// TIA Portal project "SMS-ENLAB-01-003-1501-001-PLC_V13_SP1_2_V17" (V17) (continued)
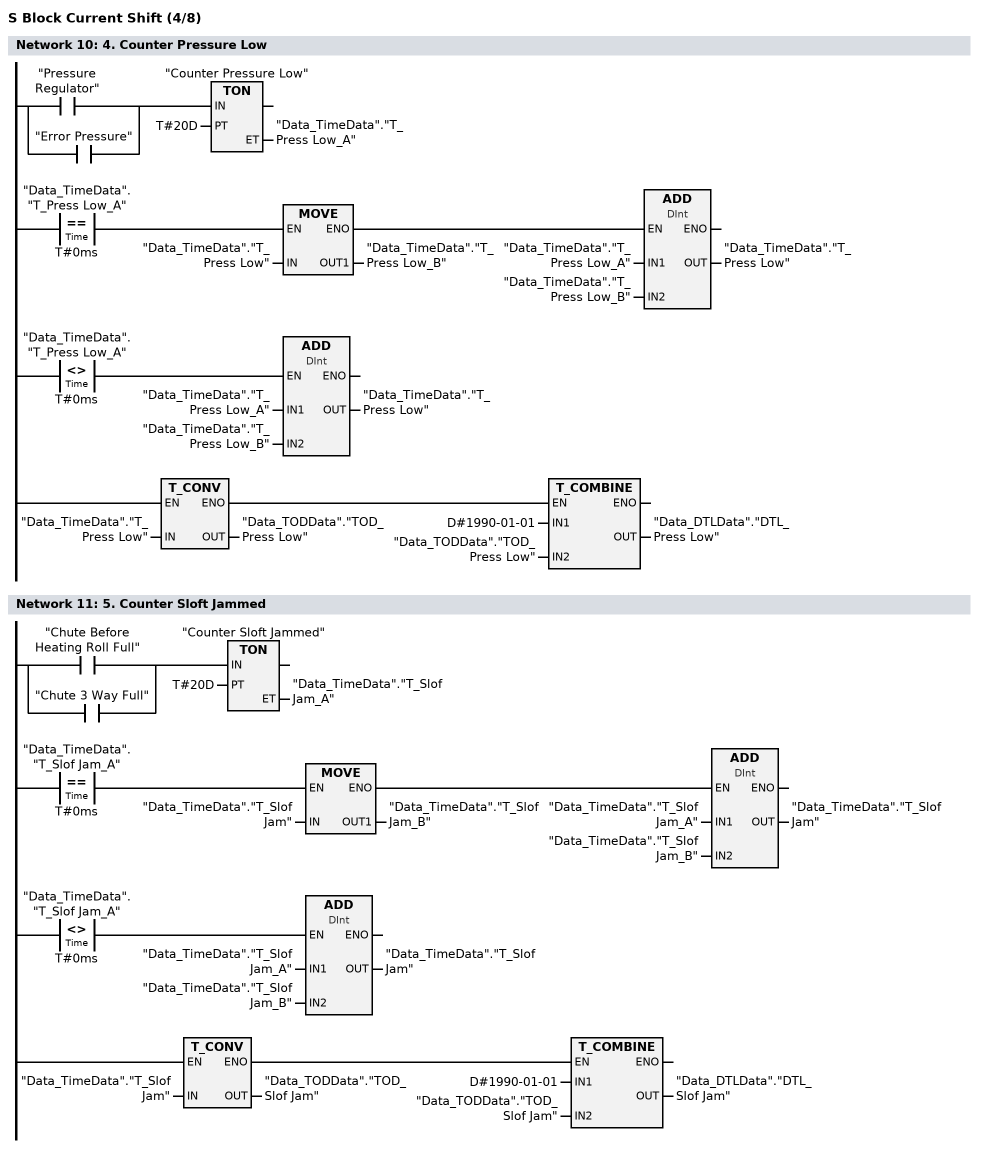
   // ENO of a box is taken as its EN; it also drops when the box reports an error
   "Counter Pressure Low".TON(IN := "Pressure Regulator" OR "Error Pressure",
                           PT := T#20D,
                           ET => "Data_TimeData"."T_Press Low_A");
   IF "Data_TimeData"."T_Press Low_A" = T#0ms THEN
       "Data_TimeData"."T_Press Low_B" := "Data_TimeData"."T_Press Low";
       "Data_TimeData"."T_Press Low" := "Data_TimeData"."T_Press Low_A" + "Data_TimeData"."T_Press Low_B";
   END_IF;
   IF "Data_TimeData"."T_Press Low_A" <> T#0ms THEN
       "Data_TimeData"."T_Press Low" := "Data_TimeData"."T_Press Low_A" + "Data_TimeData"."T_Press Low_B";
   END_IF;
   "Data_TODData"."TOD_Press Low" := T_CONV(IN := "Data_TimeData"."T_Press Low");
   "Data_DTLData"."DTL_Press Low" := T_COMBINE(IN1 := D#1990-01-01, IN2 := "Data_TODData"."TOD_Press Low");
END_REGION

REGION Network 11: 5. Counter Sloft Jammed
   // ENO of a box is taken as its EN; it also drops when the box reports an error
   "Counter Sloft Jammed".TON(IN := "Chute Before Heating Roll Full" OR "Chute 3 Way Full",
                           PT := T#20D,
                           ET => "Data_TimeData"."T_Slof Jam_A");
   IF "Data_TimeData"."T_Slof Jam_A" = T#0ms THEN
       "Data_TimeData"."T_Slof Jam_B" := "Data_TimeData"."T_Slof Jam";
       "Data_TimeData"."T_Slof Jam" := "Data_TimeData"."T_Slof Jam_A" + "Data_TimeData"."T_Slof Jam_B";
   END_IF;
   IF "Data_TimeData"."T_Slof Jam_A" <> T#0ms THEN
       "Data_TimeData"."T_Slof Jam" := "Data_TimeData"."T_Slof Jam_A" + "Data_TimeData"."T_Slof Jam_B";
   END_IF;
   "Data_TODData"."TOD_Slof Jam" := T_CONV(IN := "Data_TimeData"."T_Slof Jam");
   "Data_DTLData"."DTL_Slof Jam" := T_COMBINE(IN1 := D#1990-01-01, IN2 := "Data_TODData"."TOD_Slof Jam");
END_REGION

REGION Network 12: 7. Counter RS Pneumatic Error
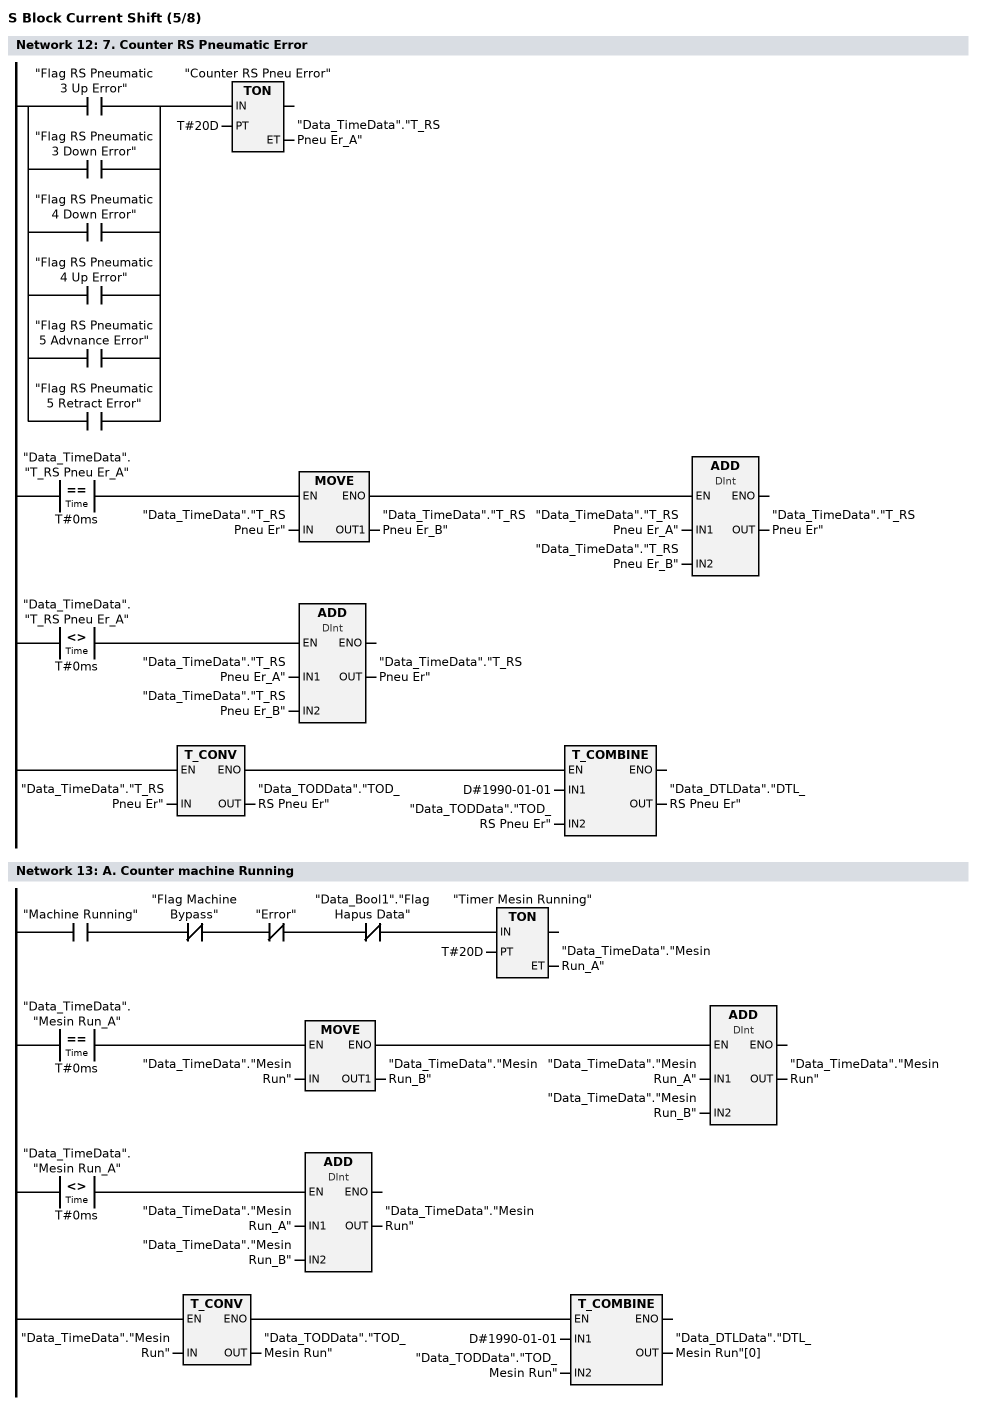
   // ENO of a box is taken as its EN; it also drops when the box reports an error
   "Counter RS Pneu Error".TON(IN := "Flag RS Pneumatic 3 Up Error" OR "Flag RS Pneumatic 3 Down Error" OR "Flag RS Pneumatic 4 Down Error" OR "Flag RS Pneumatic 4 Up Error" OR "Flag RS Pneumatic 5 Advnance Error" OR "Flag RS Pneumatic 5 Retract Error",
                           PT := T#20D,
                           ET => "Data_TimeData"."T_RS Pneu Er_A");
   IF "Data_TimeData"."T_RS Pneu Er_A" = T#0ms THEN
       "Data_TimeData"."T_RS Pneu Er_B" := "Data_TimeData"."T_RS Pneu Er";
       "Data_TimeData"."T_RS Pneu Er" := "Data_TimeData"."T_RS Pneu Er_A" + "Data_TimeData"."T_RS Pneu Er_B";
   END_IF;
   IF "Data_TimeData"."T_RS Pneu Er_A" <> T#0ms THEN
       "Data_TimeData"."T_RS Pneu Er" := "Data_TimeData"."T_RS Pneu Er_A" + "Data_TimeData"."T_RS Pneu Er_B";
   END_IF;
   "Data_TODData"."TOD_RS Pneu Er" := T_CONV(IN := "Data_TimeData"."T_RS Pneu Er");
   "Data_DTLData"."DTL_RS Pneu Er" := T_COMBINE(IN1 := D#1990-01-01, IN2 := "Data_TODData"."TOD_RS Pneu Er");
END_REGION

REGION Network 13: A. Counter machine Running
   // ENO of a box is taken as its EN; it also drops when the box reports an error
   "Timer Mesin Running".TON(IN := "Machine Running" AND NOT "Flag Machine Bypass" AND NOT "Error" AND NOT "Data_Bool1"."Flag Hapus Data",
                           PT := T#20D,
                           ET => "Data_TimeData"."Mesin Run_A");
   IF "Data_TimeData"."Mesin Run_A" = T#0ms THEN
       "Data_TimeData"."Mesin Run_B" := "Data_TimeData"."Mesin Run";
       "Data_TimeData"."Mesin Run" := "Data_TimeData"."Mesin Run_A" + "Data_TimeData"."Mesin Run_B";
   END_IF;
   IF "Data_TimeData"."Mesin Run_A" <> T#0ms THEN
       "Data_TimeData"."Mesin Run" := "Data_TimeData"."Mesin Run_A" + "Data_TimeData"."Mesin Run_B";
   END_IF;
   "Data_TODData"."TOD_Mesin Run" := T_CONV(IN := "Data_TimeData"."Mesin Run");
   "Data_DTLData"."DTL_Mesin Run"[0] := T_COMBINE(IN1 := D#1990-01-01, IN2 := "Data_TODData"."TOD_Mesin Run");
END_REGION

REGION Network 14: B. Counter machine Running Baypass Stamp
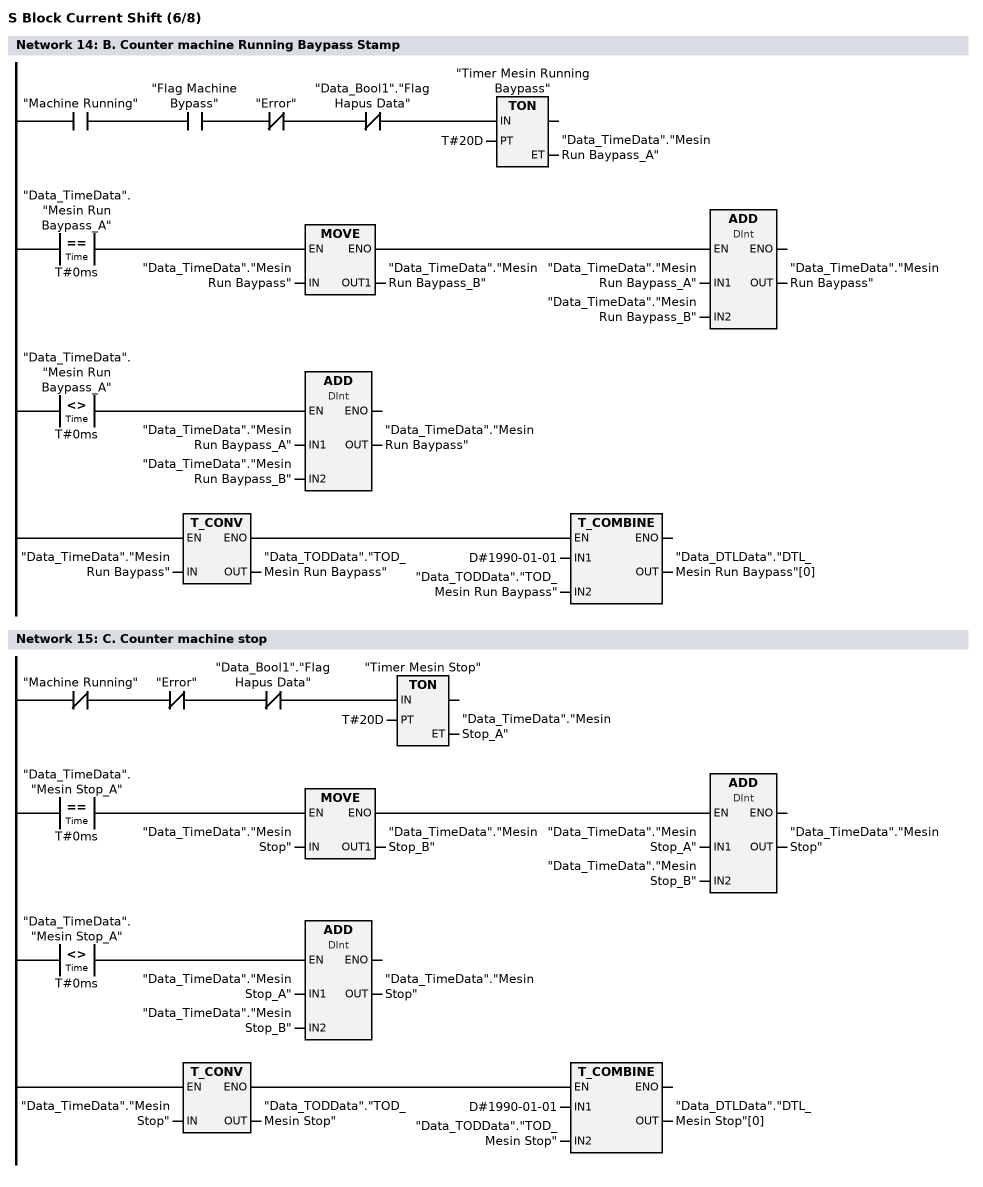
   // ENO of a box is taken as its EN; it also drops when the box reports an error
   "Timer Mesin Running Baypass".TON(IN := "Machine Running" AND "Flag Machine Bypass" AND NOT "Error" AND NOT "Data_Bool1"."Flag Hapus Data",
                           PT := T#20D,
                           ET => "Data_TimeData"."Mesin Run Baypass_A");
   IF "Data_TimeData"."Mesin Run Baypass_A" = T#0ms THEN
       "Data_TimeData"."Mesin Run Baypass_B" := "Data_TimeData"."Mesin Run Baypass";
       "Data_TimeData"."Mesin Run Baypass" := "Data_TimeData"."Mesin Run Baypass_A" + "Data_TimeData"."Mesin Run Baypass_B";
   END_IF;
   IF "Data_TimeData"."Mesin Run Baypass_A" <> T#0ms THEN
       "Data_TimeData"."Mesin Run Baypass" := "Data_TimeData"."Mesin Run Baypass_A" + "Data_TimeData"."Mesin Run Baypass_B";
   END_IF;
   "Data_TODData"."TOD_Mesin Run Baypass" := T_CONV(IN := "Data_TimeData"."Mesin Run Baypass");
   "Data_DTLData"."DTL_Mesin Run Baypass"[0] := T_COMBINE(IN1 := D#1990-01-01,
                           IN2 := "Data_TODData"."TOD_Mesin Run Baypass");
END_REGION

REGION Network 15: C. Counter machine stop
   // ENO of a box is taken as its EN; it also drops when the box reports an error
   "Timer Mesin Stop".TON(IN := NOT "Machine Running" AND NOT "Error" AND NOT "Data_Bool1"."Flag Hapus Data",
                          PT := T#20D,
                          ET => "Data_TimeData"."Mesin Stop_A");
   IF "Data_TimeData"."Mesin Stop_A" = T#0ms THEN
       "Data_TimeData"."Mesin Stop_B" := "Data_TimeData"."Mesin Stop";
       "Data_TimeData"."Mesin Stop" := "Data_TimeData"."Mesin Stop_A" + "Data_TimeData"."Mesin Stop_B";
   END_IF;
   IF "Data_TimeData"."Mesin Stop_A" <> T#0ms THEN
       "Data_TimeData"."Mesin Stop" := "Data_TimeData"."Mesin Stop_A" + "Data_TimeData"."Mesin Stop_B";
   END_IF;
   "Data_TODData"."TOD_Mesin Stop" := T_CONV(IN := "Data_TimeData"."Mesin Stop");
   "Data_DTLData"."DTL_Mesin Stop"[0] := T_COMBINE(IN1 := D#1990-01-01, IN2 := "Data_TODData"."TOD_Mesin Stop");
END_REGION

REGION Network 16: D. Counter Machine Error
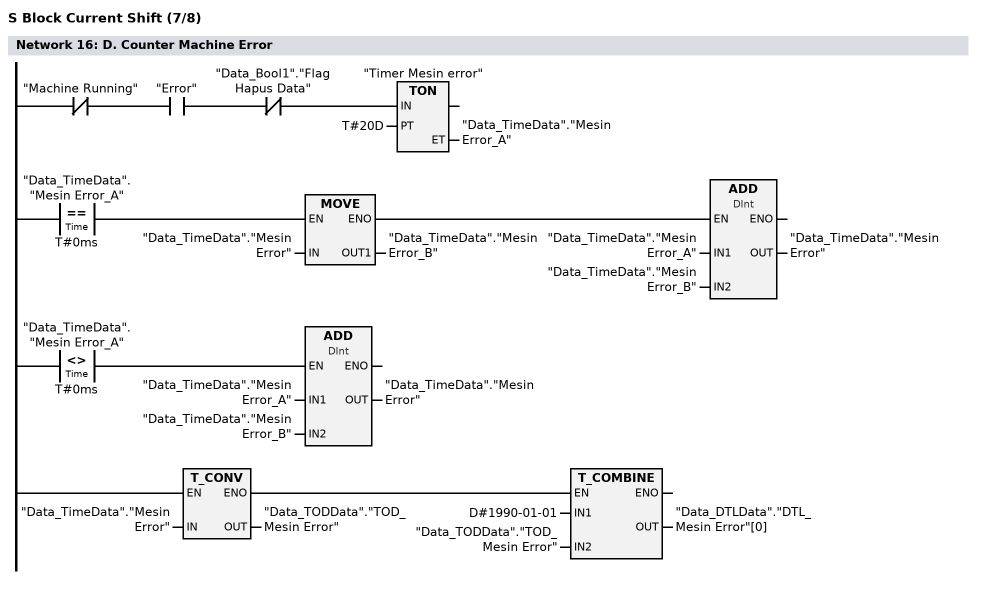
   // ENO of a box is taken as its EN; it also drops when the box reports an error
   "Timer Mesin error".TON(IN := NOT "Machine Running" AND "Error" AND NOT "Data_Bool1"."Flag Hapus Data",
                           PT := T#20D,
                           ET => "Data_TimeData"."Mesin Error_A");
   IF "Data_TimeData"."Mesin Error_A" = T#0ms THEN
       "Data_TimeData"."Mesin Error_B" := "Data_TimeData"."Mesin Error";
       "Data_TimeData"."Mesin Error" := "Data_TimeData"."Mesin Error_A" + "Data_TimeData"."Mesin Error_B";
   END_IF;
   IF "Data_TimeData"."Mesin Error_A" <> T#0ms THEN
       "Data_TimeData"."Mesin Error" := "Data_TimeData"."Mesin Error_A" + "Data_TimeData"."Mesin Error_B";
   END_IF;
   "Data_TODData"."TOD_Mesin Error" := T_CONV(IN := "Data_TimeData"."Mesin Error");
   "Data_DTLData"."DTL_Mesin Error"[0] := T_COMBINE(IN1 := D#1990-01-01,
                           IN2 := "Data_TODData"."TOD_Mesin Error");
END_REGION

REGION Network 17: % Persen Counter Mesin Terhadap Lama Current Shift
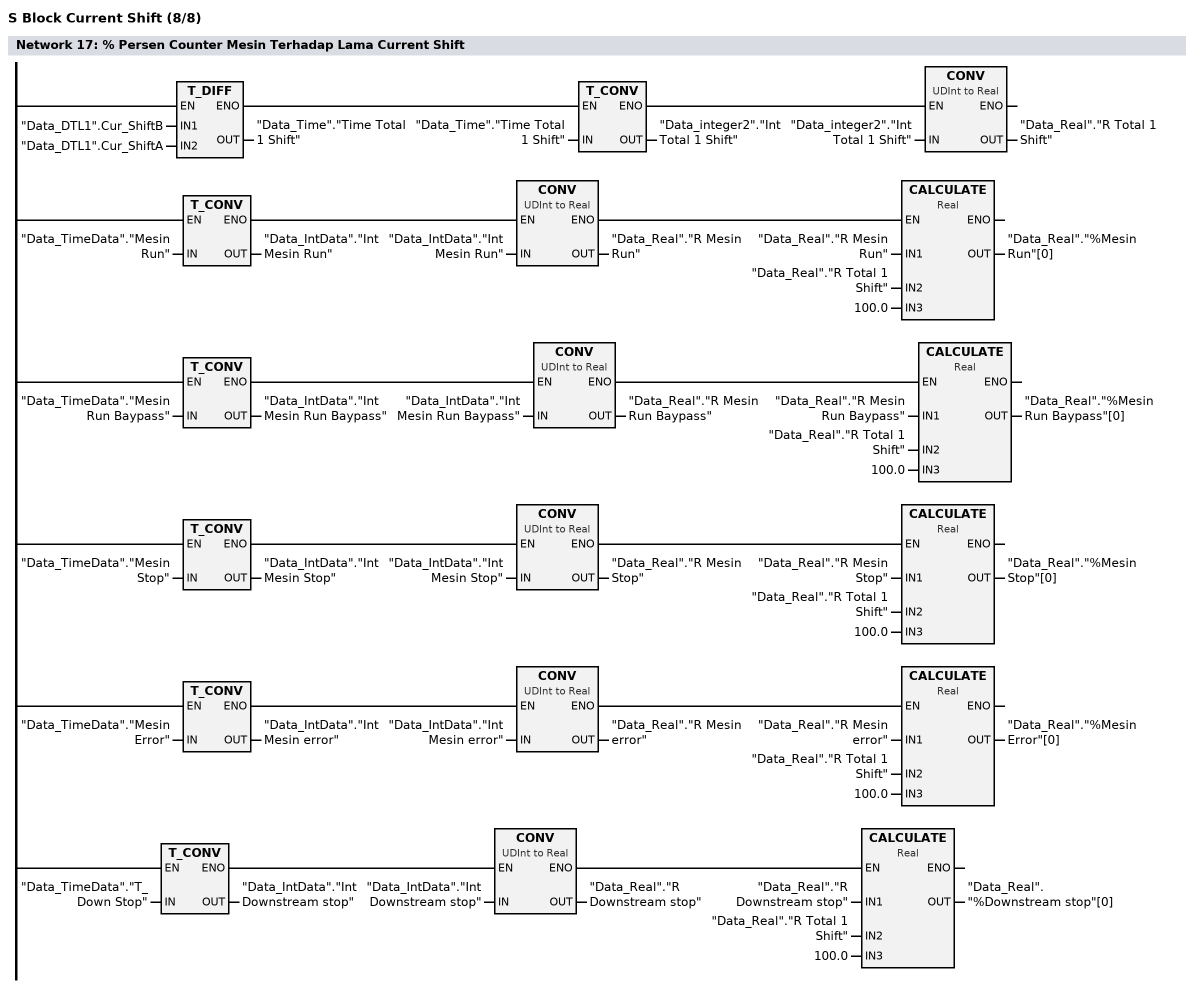
   // ENO of a box is taken as its EN; it also drops when the box reports an error
   "Data_Time"."Time Total 1 Shift" := T_DIFF(IN1 := "Data_DTL1".Cur_ShiftB, IN2 := "Data_DTL1".Cur_ShiftA);
   "Data_integer2"."Int Total 1 Shift" := T_CONV(IN := "Data_Time"."Time Total 1 Shift");
   "Data_Real"."R Total 1 Shift" := UDINT_TO_REAL("Data_integer2"."Int Total 1 Shift");
   "Data_IntData"."Int Mesin Run" := T_CONV(IN := "Data_TimeData"."Mesin Run");
   "Data_Real"."R Mesin Run" := UDINT_TO_REAL("Data_IntData"."Int Mesin Run");
   "Data_Real"."%Mesin Run"[0] := ("Data_Real"."R Mesin Run"/"Data_Real"."R Total 1 Shift")*100.0;
   "Data_IntData"."Int Mesin Run Baypass" := T_CONV(IN := "Data_TimeData"."Mesin Run Baypass");
   "Data_Real"."R Mesin Run Baypass" := UDINT_TO_REAL("Data_IntData"."Int Mesin Run Baypass");
   "Data_Real"."%Mesin Run Baypass"[0] := ("Data_Real"."R Mesin Run Baypass"/"Data_Real"."R Total 1 Shift")*100.0;
   "Data_IntData"."Int Mesin Stop" := T_CONV(IN := "Data_TimeData"."Mesin Stop");
   "Data_Real"."R Mesin Stop" := UDINT_TO_REAL("Data_IntData"."Int Mesin Stop");
   "Data_Real"."%Mesin Stop"[0] := ("Data_Real"."R Mesin Stop"/"Data_Real"."R Total 1 Shift")*100.0;
   "Data_IntData"."Int Mesin error" := T_CONV(IN := "Data_TimeData"."Mesin Error");
   "Data_Real"."R Mesin error" := UDINT_TO_REAL("Data_IntData"."Int Mesin error");
   "Data_Real"."%Mesin Error"[0] := ("Data_Real"."R Mesin error"/"Data_Real"."R Total 1 Shift")*100.0;
   "Data_IntData"."Int Downstream stop" := T_CONV(IN := "Data_TimeData"."T_Down Stop");
   "Data_Real"."R Downstream stop" := UDINT_TO_REAL("Data_IntData"."Int Downstream stop");
   "Data_Real"."%Downstream stop"[0] := ("Data_Real"."R Downstream stop"/"Data_Real"."R Total 1 Shift")*100.0;
END_REGION
END_FUNCTION_BLOCK

FUNCTION_BLOCK "Block Labeling"   // FB5, LAD
{ S7_Optimized_Access := 'TRUE' }
VERSION : 0.1
   VAR_TEMP   // added for the SCL form of the ladder/FBD networks
      _w1 : Bool;
      _w2 : Bool;
      _w3 : Bool;
      _w4 : Bool;
      _w5 : Bool;
   END_VAR
BEGIN

REGION Network 1: By pass ON
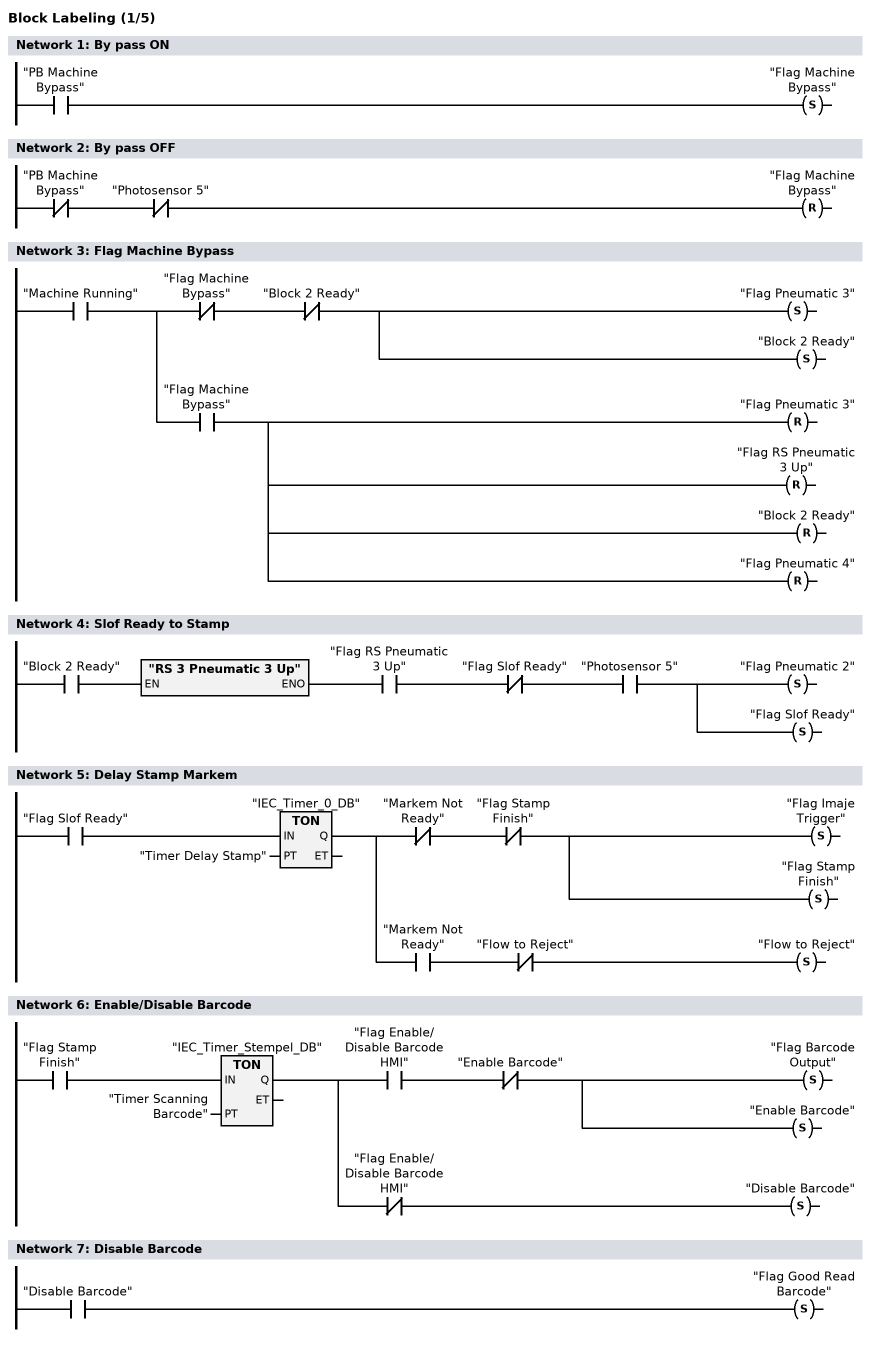
   RUNG wire#powerrail
      Contact( "PB Machine Bypass" )
      S_Coil( "Flag Machine Bypass" )
   END_RUNG
   // the same network as SCL:
   IF "PB Machine Bypass" THEN "Flag Machine Bypass" := TRUE; END_IF;
END_REGION

REGION Network 2: By pass OFF
   RUNG wire#powerrail
      I_Contact( "PB Machine Bypass" )
      I_Contact( "Photosensor 5" )
      R_Coil( "Flag Machine Bypass" )
   END_RUNG
   // the same network as SCL:
   IF NOT "PB Machine Bypass" AND NOT "Photosensor 5" THEN "Flag Machine Bypass" := FALSE; END_IF;
END_REGION

REGION Network 3: Flag Machine Bypass
   RUNG wire#powerrail
      Contact( "Machine Running" )
      wire#w1
      I_Contact( "Flag Machine Bypass" )
      I_Contact( "Block 2 Ready" )
      wire#w2
      S_Coil( "Flag Pneumatic 3" )
   END_RUNG
   RUNG wire#w2
      S_Coil( "Block 2 Ready" )
   END_RUNG
   RUNG wire#w1
      Contact( "Flag Machine Bypass" )
      wire#w3
      R_Coil( "Flag Pneumatic 3" )
   END_RUNG
   RUNG wire#w3
      R_Coil( "Flag RS Pneumatic 3 Up" )
   END_RUNG
   RUNG wire#w3
      R_Coil( "Block 2 Ready" )
   END_RUNG
   RUNG wire#w3
      R_Coil( "Flag Pneumatic 4" )
   END_RUNG
   // the same network as SCL:
   IF "Machine Running" AND NOT "Flag Machine Bypass" AND NOT "Block 2 Ready" THEN
       "Flag Pneumatic 3" := TRUE;
       "Block 2 Ready" := TRUE;
   END_IF;
   IF "Machine Running" AND "Flag Machine Bypass" THEN
       "Flag Pneumatic 3" := FALSE;
       "Flag RS Pneumatic 3 Up" := FALSE;
       "Block 2 Ready" := FALSE;
       "Flag Pneumatic 4" := FALSE;
   END_IF;
END_REGION

REGION Network 4: Slof Ready to Stamp
   RUNG wire#powerrail
      Contact( "Block 2 Ready" )
      "RS 3 Pneumatic 3 Up"()
      Contact( "Flag RS Pneumatic 3 Up" )
      I_Contact( "Flag Slof Ready" )
      Contact( "Photosensor 5" )
      wire#w1
      S_Coil( "Flag Pneumatic 2" )
   END_RUNG
   RUNG wire#w1
      S_Coil( "Flag Slof Ready" )
   END_RUNG
   // the same network as SCL:
   "RS 3 Pneumatic 3 Up"(EN := "Block 2 Ready", ENO => #_w1);
   IF #_w1 AND "Flag RS Pneumatic 3 Up" AND NOT "Flag Slof Ready" AND "Photosensor 5" THEN
       "Flag Pneumatic 2" := TRUE;
       "Flag Slof Ready" := TRUE;
   END_IF;
END_REGION

REGION Network 5: Delay Stamp Markem
   "IEC_Timer_0_DB".TON(IN := "Flag Slof Ready", PT := "Timer Delay Stamp");
   IF "IEC_Timer_0_DB".Q AND NOT "Markem Not Ready" AND NOT "Flag Stamp Finish" THEN
       "Flag Imaje Trigger" := TRUE;
       "Flag Stamp Finish" := TRUE;
   END_IF;
   IF "IEC_Timer_0_DB".Q AND "Markem Not Ready" AND NOT "Flow to Reject" THEN
       "Flow to Reject" := TRUE;
   END_IF;
END_REGION

REGION Network 6: Enable/Disable Barcode
   "IEC_Timer_Stempel_DB".TON(IN := "Flag Stamp Finish", PT := "Timer Scanning Barcode");
   IF "IEC_Timer_Stempel_DB".Q AND "Flag Enable/Disable Barcode HMI" AND NOT "Enable Barcode" THEN
       "Flag Barcode Output" := TRUE;
       "Enable Barcode" := TRUE;
   END_IF;
   IF "IEC_Timer_Stempel_DB".Q AND NOT "Flag Enable/Disable Barcode HMI" THEN
       "Disable Barcode" := TRUE;
   END_IF;
END_REGION

REGION Network 7: Disable Barcode
   RUNG wire#powerrail
      Contact( "Disable Barcode" )
      S_Coil( "Flag Good Read Barcode" )
   END_RUNG
   // the same network as SCL:
   IF "Disable Barcode" THEN "Flag Good Read Barcode" := TRUE; END_IF;
END_REGION

REGION Network 8: Check Barcode
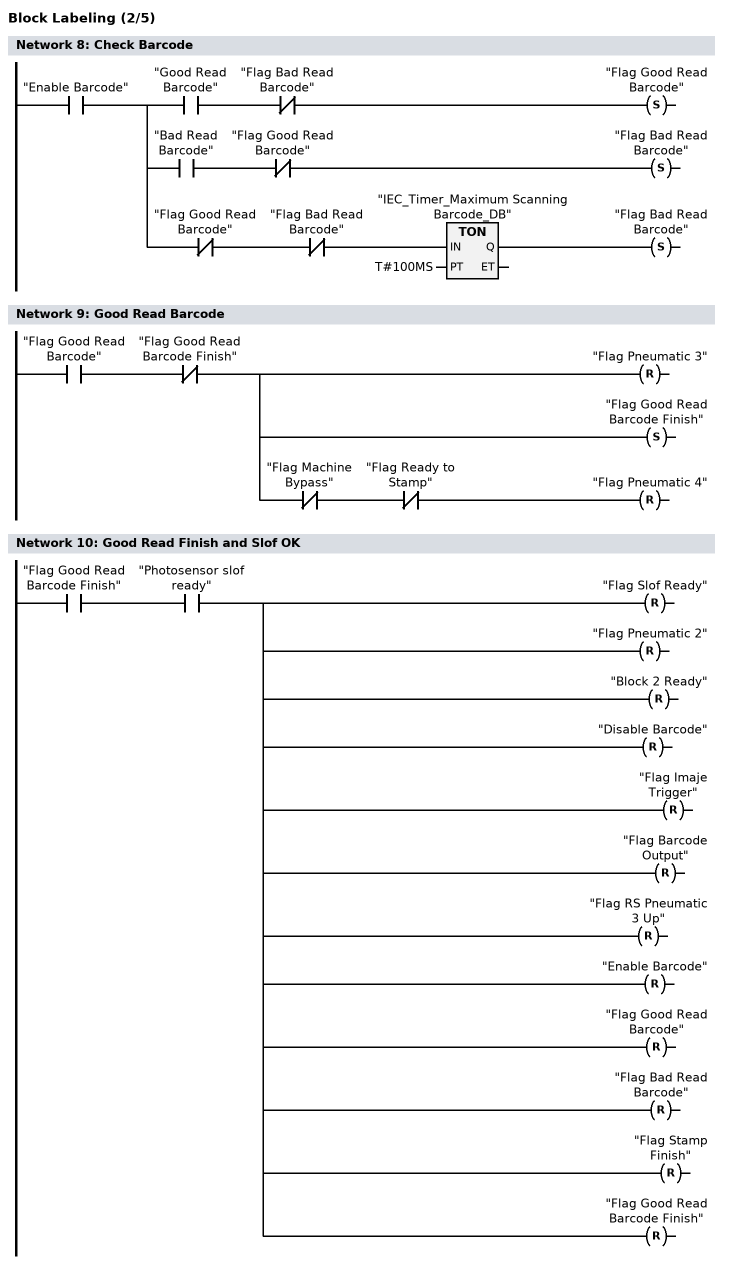
   IF "Enable Barcode" AND "Good Read Barcode" AND NOT "Flag Bad Read Barcode" THEN
       "Flag Good Read Barcode" := TRUE;
   END_IF;
   IF "Enable Barcode" AND "Bad Read Barcode" AND NOT "Flag Good Read Barcode" THEN
       "Flag Bad Read Barcode" := TRUE;
   END_IF;
   "IEC_Timer_Maximum Scanning Barcode_DB".TON(IN := "Enable Barcode" AND NOT "Flag Good Read Barcode" AND NOT "Flag Bad Read Barcode",
                           PT := T#100MS);
   IF "IEC_Timer_Maximum Scanning Barcode_DB".Q THEN "Flag Bad Read Barcode" := TRUE; END_IF;
END_REGION

REGION Network 9: Good Read Barcode
   RUNG wire#powerrail
      Contact( "Flag Good Read Barcode" )
      I_Contact( "Flag Good Read Barcode Finish" )
      wire#w1
      R_Coil( "Flag Pneumatic 3" )
   END_RUNG
   RUNG wire#w1
      S_Coil( "Flag Good Read Barcode Finish" )
   END_RUNG
   RUNG wire#w1
      I_Contact( "Flag Machine Bypass" )
      I_Contact( "Flag Ready to Stamp" )
      R_Coil( "Flag Pneumatic 4" )
   END_RUNG
   // the same network as SCL:
   #_w1 := "Flag Good Read Barcode" AND NOT "Flag Good Read Barcode Finish";
   IF #_w1 THEN
       "Flag Pneumatic 3" := FALSE;
       "Flag Good Read Barcode Finish" := TRUE;
   END_IF;
   IF #_w1 AND NOT "Flag Machine Bypass" AND NOT "Flag Ready to Stamp" THEN
       "Flag Pneumatic 4" := FALSE;
   END_IF;
END_REGION

REGION Network 10: Good Read Finish and Slof OK
   RUNG wire#powerrail
      Contact( "Flag Good Read Barcode Finish" )
      Contact( "Photosensor slof ready" )
      wire#w1
      R_Coil( "Flag Slof Ready" )
   END_RUNG
   RUNG wire#w1
      R_Coil( "Flag Pneumatic 2" )
   END_RUNG
   RUNG wire#w1
      R_Coil( "Block 2 Ready" )
   END_RUNG
   RUNG wire#w1
      R_Coil( "Disable Barcode" )
   END_RUNG
   RUNG wire#w1
      R_Coil( "Flag Imaje Trigger" )
   END_RUNG
   RUNG wire#w1
      R_Coil( "Flag Barcode Output" )
   END_RUNG
   RUNG wire#w1
      R_Coil( "Flag RS Pneumatic 3 Up" )
   END_RUNG
   RUNG wire#w1
      R_Coil( "Enable Barcode" )
   END_RUNG
   RUNG wire#w1
      R_Coil( "Flag Good Read Barcode" )
   END_RUNG
   RUNG wire#w1
      R_Coil( "Flag Bad Read Barcode" )
   END_RUNG
   RUNG wire#w1
      R_Coil( "Flag Stamp Finish" )
   END_RUNG
   RUNG wire#w1
      R_Coil( "Flag Good Read Barcode Finish" )
   END_RUNG
   // the same network as SCL:
   IF "Flag Good Read Barcode Finish" AND "Photosensor slof ready" THEN
       "Flag Slof Ready" := FALSE;
       "Flag Pneumatic 2" := FALSE;
       "Block 2 Ready" := FALSE;
       "Disable Barcode" := FALSE;
       "Flag Imaje Trigger" := FALSE;
       "Flag Barcode Output" := FALSE;
       "Flag RS Pneumatic 3 Up" := FALSE;
       "Enable Barcode" := FALSE;
       "Flag Good Read Barcode" := FALSE;
       "Flag Bad Read Barcode" := FALSE;
       "Flag Stamp Finish" := FALSE;
       "Flag Good Read Barcode Finish" := FALSE;
   END_IF;
END_REGION

REGION Network 11: Set Section Reject
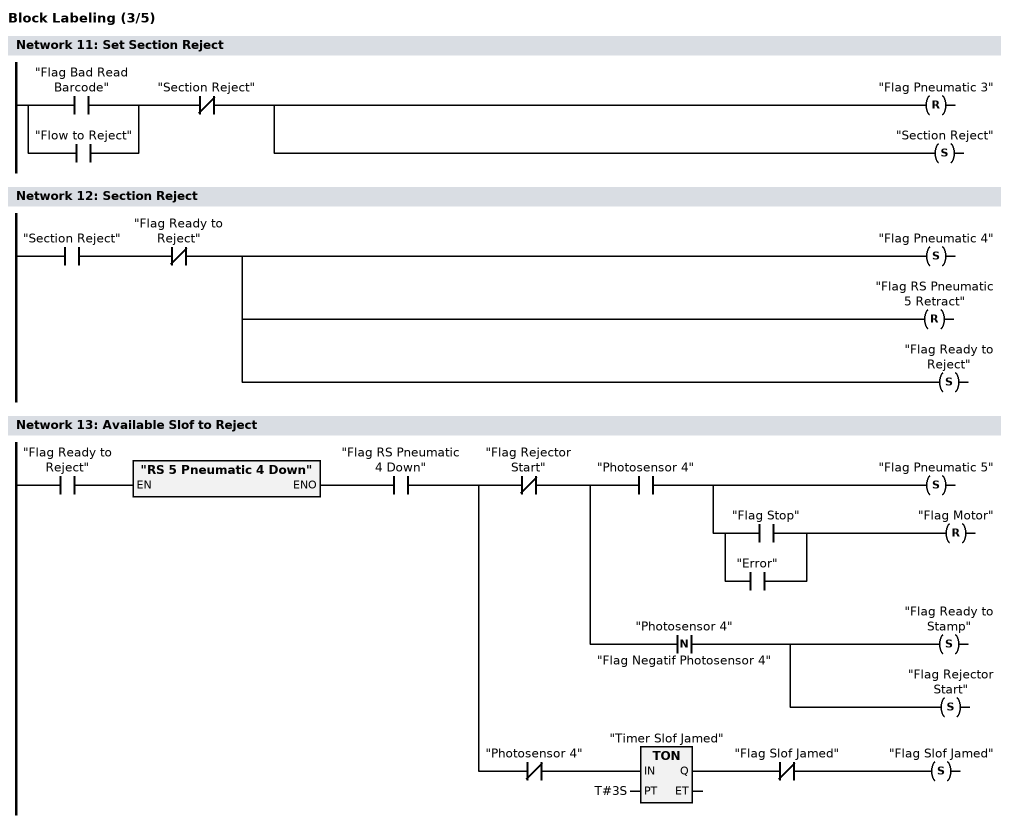
   RUNG wire#powerrail
      Contact( "Flag Bad Read Barcode" )
      wire#w1
      I_Contact( "Section Reject" )
      wire#w2
      R_Coil( "Flag Pneumatic 3" )
   END_RUNG
   RUNG wire#powerrail
      Contact( "Flow to Reject" )
   END_RUNG wire#w1
   RUNG wire#w2
      S_Coil( "Section Reject" )
   END_RUNG
   // the same network as SCL:
   IF ("Flag Bad Read Barcode" OR "Flow to Reject") AND NOT "Section Reject" THEN
       "Flag Pneumatic 3" := FALSE;
       "Section Reject" := TRUE;
   END_IF;
END_REGION

REGION Network 12: Section Reject
   RUNG wire#powerrail
      Contact( "Section Reject" )
      I_Contact( "Flag Ready to Reject" )
      wire#w1
      S_Coil( "Flag Pneumatic 4" )
   END_RUNG
   RUNG wire#w1
      R_Coil( "Flag RS Pneumatic 5 Retract" )
   END_RUNG
   RUNG wire#w1
      S_Coil( "Flag Ready to Reject" )
   END_RUNG
   // the same network as SCL:
   IF "Section Reject" AND NOT "Flag Ready to Reject" THEN
       "Flag Pneumatic 4" := TRUE;
       "Flag RS Pneumatic 5 Retract" := FALSE;
       "Flag Ready to Reject" := TRUE;
   END_IF;
END_REGION

REGION Network 13: Available Slof to Reject
   "RS 5 Pneumatic 4 Down"(EN := "Flag Ready to Reject", ENO => #_w1);
   #_w2 := #_w1 AND "Flag RS Pneumatic 4 Down";
   #_w3 := #_w2 AND NOT "Flag Rejector Start";
   #_w4 := #_w3 AND "Photosensor 4";
   IF #_w4 THEN "Flag Pneumatic 5" := TRUE; END_IF;
   IF #_w4 AND ("Flag Stop" OR "Error") THEN "Flag Motor" := FALSE; END_IF;
   #_w5 := #_w3 AND NOT "Photosensor 4" AND "Flag Negatif Photosensor 4";   // falling edge of "Photosensor 4"
   "Flag Negatif Photosensor 4" := "Photosensor 4";
   IF #_w5 THEN
       "Flag Ready to Stamp" := TRUE;
       "Flag Rejector Start" := TRUE;
   END_IF;
   "Timer Slof Jamed".TON(IN := #_w2 AND NOT "Photosensor 4", PT := T#3S);
   IF "Timer Slof Jamed".Q AND NOT "Flag Slof Jamed" THEN "Flag Slof Jamed" := TRUE; END_IF;
END_REGION

REGION Network 14: Ready to Stamp again
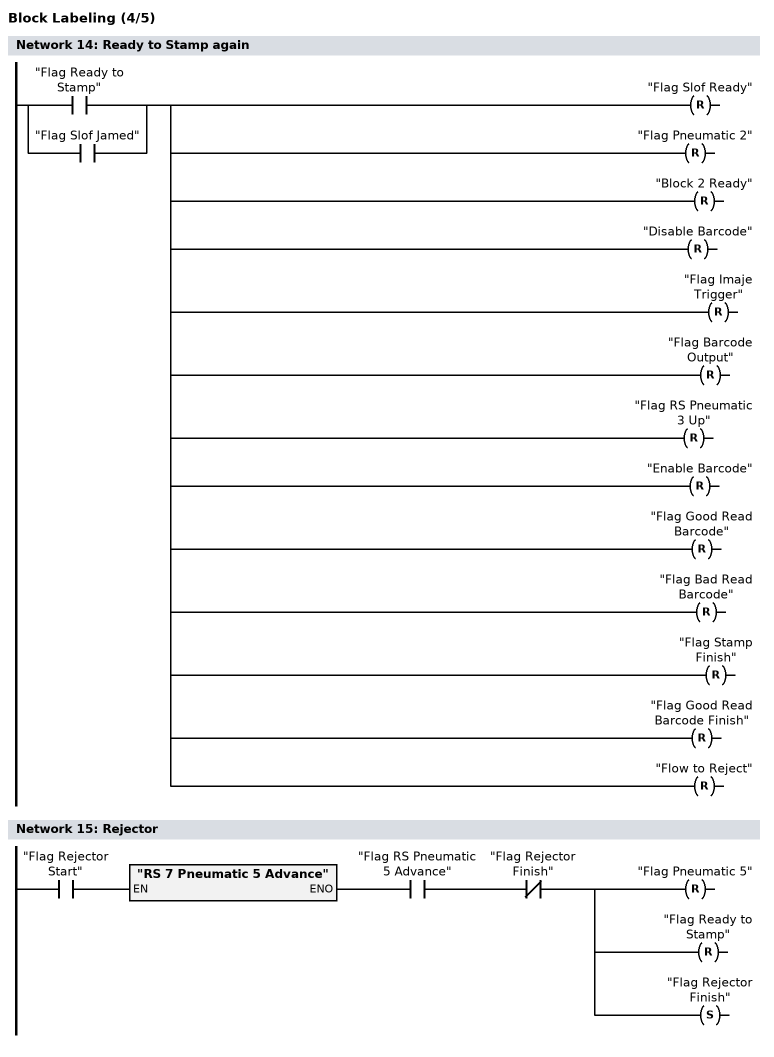
   RUNG wire#powerrail
      Contact( "Flag Ready to Stamp" )
      wire#w1
      R_Coil( "Flag Slof Ready" )
   END_RUNG
   RUNG wire#powerrail
      Contact( "Flag Slof Jamed" )
   END_RUNG wire#w1
   RUNG wire#w1
      R_Coil( "Flag Pneumatic 2" )
   END_RUNG
   RUNG wire#w1
      R_Coil( "Block 2 Ready" )
   END_RUNG
   RUNG wire#w1
      R_Coil( "Disable Barcode" )
   END_RUNG
   RUNG wire#w1
      R_Coil( "Flag Imaje Trigger" )
   END_RUNG
   RUNG wire#w1
      R_Coil( "Flag Barcode Output" )
   END_RUNG
   RUNG wire#w1
      R_Coil( "Flag RS Pneumatic 3 Up" )
   END_RUNG
   RUNG wire#w1
      R_Coil( "Enable Barcode" )
   END_RUNG
   RUNG wire#w1
      R_Coil( "Flag Good Read Barcode" )
   END_RUNG
   RUNG wire#w1
      R_Coil( "Flag Bad Read Barcode" )
   END_RUNG
   RUNG wire#w1
      R_Coil( "Flag Stamp Finish" )
   END_RUNG
   RUNG wire#w1
      R_Coil( "Flag Good Read Barcode Finish" )
   END_RUNG
   RUNG wire#w1
      R_Coil( "Flow to Reject" )
   END_RUNG
   // the same network as SCL:
   IF "Flag Ready to Stamp" OR "Flag Slof Jamed" THEN
       "Flag Slof Ready" := FALSE;
       "Flag Pneumatic 2" := FALSE;
       "Block 2 Ready" := FALSE;
       "Disable Barcode" := FALSE;
       "Flag Imaje Trigger" := FALSE;
       "Flag Barcode Output" := FALSE;
       "Flag RS Pneumatic 3 Up" := FALSE;
       "Enable Barcode" := FALSE;
       "Flag Good Read Barcode" := FALSE;
       "Flag Bad Read Barcode" := FALSE;
       "Flag Stamp Finish" := FALSE;
       "Flag Good Read Barcode Finish" := FALSE;
       "Flow to Reject" := FALSE;
   END_IF;
END_REGION

REGION Network 15: Rejector
   RUNG wire#powerrail
      Contact( "Flag Rejector Start" )
      "RS 7 Pneumatic 5 Advance"()
      Contact( "Flag RS Pneumatic 5 Advance" )
      I_Contact( "Flag Rejector Finish" )
      wire#w1
      R_Coil( "Flag Pneumatic 5" )
   END_RUNG
   RUNG wire#w1
      R_Coil( "Flag Ready to Stamp" )
   END_RUNG
   RUNG wire#w1
      S_Coil( "Flag Rejector Finish" )
   END_RUNG
   // the same network as SCL:
   "RS 7 Pneumatic 5 Advance"(EN := "Flag Rejector Start", ENO => #_w1);
   IF #_w1 AND "Flag RS Pneumatic 5 Advance" AND NOT "Flag Rejector Finish" THEN
       "Flag Pneumatic 5" := FALSE;
       "Flag Ready to Stamp" := FALSE;
       "Flag Rejector Finish" := TRUE;
   END_IF;
END_REGION

REGION Network 16: Rejector Finish
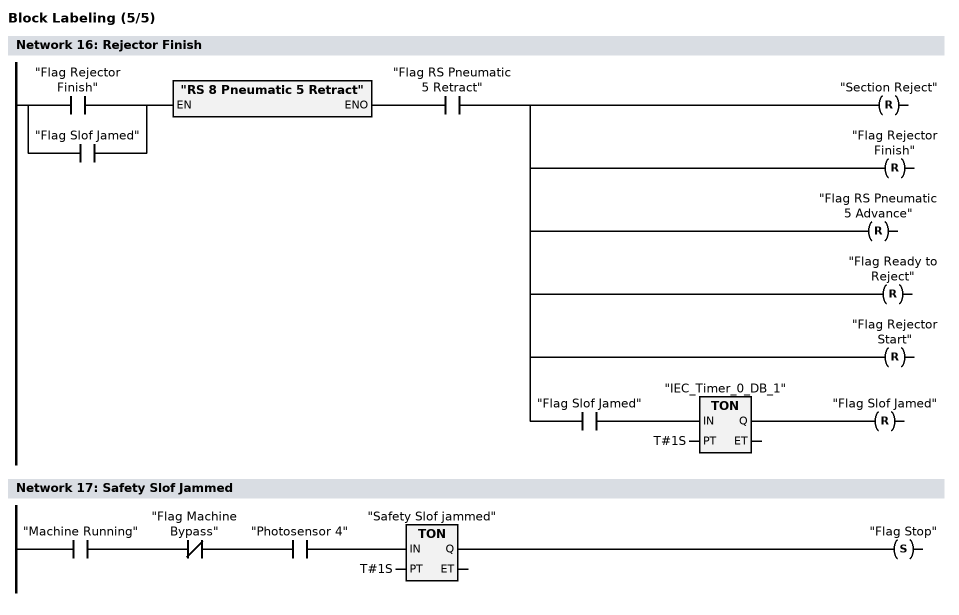
   "RS 8 Pneumatic 5 Retract"(EN := "Flag Rejector Finish" OR "Flag Slof Jamed", ENO => #_w1);
   #_w2 := #_w1 AND "Flag RS Pneumatic 5 Retract";
   IF #_w2 THEN
       "Section Reject" := FALSE;
       "Flag Rejector Finish" := FALSE;
       "Flag RS Pneumatic 5 Advance" := FALSE;
       "Flag Ready to Reject" := FALSE;
       "Flag Rejector Start" := FALSE;
   END_IF;
   "IEC_Timer_0_DB_1".TON(IN := #_w2 AND "Flag Slof Jamed", PT := T#1S);
   IF "IEC_Timer_0_DB_1".Q THEN "Flag Slof Jamed" := FALSE; END_IF;
END_REGION

REGION Network 17: Safety Slof Jammed
   "Safety Slof jammed".TON(IN := "Machine Running" AND NOT "Flag Machine Bypass" AND "Photosensor 4",
                           PT := T#1S);
   IF "Safety Slof jammed".Q THEN "Flag Stop" := TRUE; END_IF;
END_REGION
END_FUNCTION_BLOCK

FUNCTION_BLOCK "Block Focke"   // FB6, LAD
{ S7_Optimized_Access := 'TRUE' }
VERSION : 0.1
   VAR_TEMP   // added for the SCL form of the ladder/FBD networks
      _w1 : Bool;
   END_VAR
BEGIN

REGION Network 1: Enable/Disable Error Chute Before Heating Roll
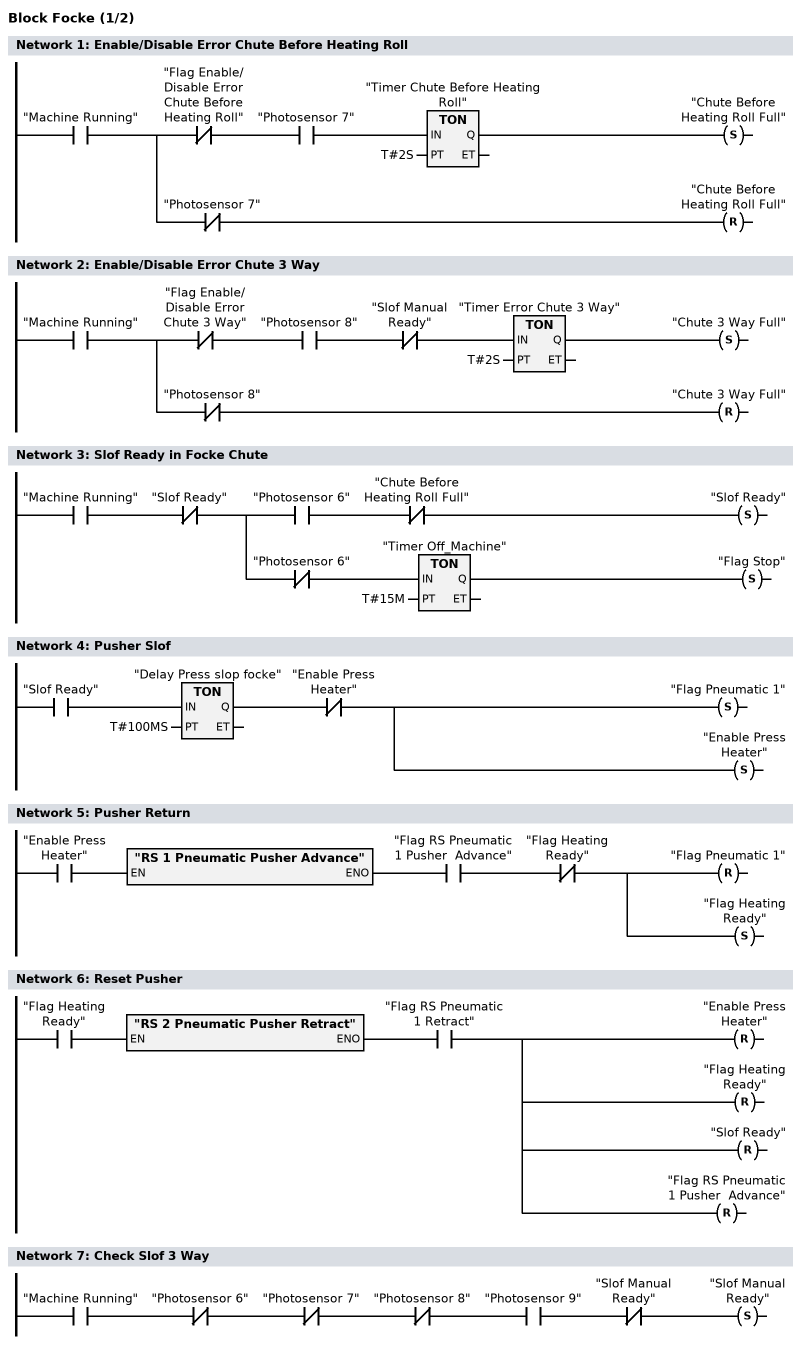
   "Timer Chute Before Heating Roll".TON(IN := "Machine Running" AND NOT "Flag Enable/Disable Error Chute Before Heating Roll" AND "Photosensor 7",
                           PT := T#2S);
   IF "Timer Chute Before Heating Roll".Q THEN "Chute Before Heating Roll Full" := TRUE; END_IF;
   IF "Machine Running" AND NOT "Photosensor 7" THEN "Chute Before Heating Roll Full" := FALSE; END_IF;
END_REGION

REGION Network 2: Enable/Disable Error Chute 3 Way
   "Timer Error Chute 3 Way".TON(IN := "Machine Running" AND NOT "Flag Enable/Disable Error Chute 3 Way" AND "Photosensor 8" AND NOT "Slof Manual Ready",
                           PT := T#2S);
   IF "Timer Error Chute 3 Way".Q THEN "Chute 3 Way Full" := TRUE; END_IF;
   IF "Machine Running" AND NOT "Photosensor 8" THEN "Chute 3 Way Full" := FALSE; END_IF;
END_REGION

REGION Network 3: Slof Ready in Focke Chute
   #_w1 := "Machine Running" AND NOT "Slof Ready";
   IF #_w1 AND "Photosensor 6" AND NOT "Chute Before Heating Roll Full" THEN "Slof Ready" := TRUE; END_IF;
   "Timer Off_Machine".TON(IN := #_w1 AND NOT "Photosensor 6", PT := T#15M);
   IF "Timer Off_Machine".Q THEN "Flag Stop" := TRUE; END_IF;
END_REGION

REGION Network 4: Pusher Slof
   "Delay Press slop focke".TON(IN := "Slof Ready", PT := T#100MS);
   IF "Delay Press slop focke".Q AND NOT "Enable Press Heater" THEN
       "Flag Pneumatic 1" := TRUE;
       "Enable Press Heater" := TRUE;
   END_IF;
END_REGION

REGION Network 5: Pusher Return
   RUNG wire#powerrail
      Contact( "Enable Press Heater" )
      "RS 1 Pneumatic Pusher Advance"()
      Contact( "Flag RS Pneumatic 1 Pusher  Advance" )
      I_Contact( "Flag Heating Ready" )
      wire#w1
      R_Coil( "Flag Pneumatic 1" )
   END_RUNG
   RUNG wire#w1
      S_Coil( "Flag Heating Ready" )
   END_RUNG
   // the same network as SCL:
   "RS 1 Pneumatic Pusher Advance"(EN := "Enable Press Heater", ENO => #_w1);
   IF #_w1 AND "Flag RS Pneumatic 1 Pusher  Advance" AND NOT "Flag Heating Ready" THEN
       "Flag Pneumatic 1" := FALSE;
       "Flag Heating Ready" := TRUE;
   END_IF;
END_REGION

REGION Network 6: Reset Pusher
   RUNG wire#powerrail
      Contact( "Flag Heating Ready" )
      "RS 2 Pneumatic Pusher Retract"()
      Contact( "Flag RS Pneumatic 1 Retract" )
      wire#w1
      R_Coil( "Enable Press Heater" )
   END_RUNG
   RUNG wire#w1
      R_Coil( "Flag Heating Ready" )
   END_RUNG
   RUNG wire#w1
      R_Coil( "Slof Ready" )
   END_RUNG
   RUNG wire#w1
      R_Coil( "Flag RS Pneumatic 1 Pusher  Advance" )
   END_RUNG
   // the same network as SCL:
   "RS 2 Pneumatic Pusher Retract"(EN := "Flag Heating Ready", ENO => #_w1);
   IF #_w1 AND "Flag RS Pneumatic 1 Retract" THEN
       "Enable Press Heater" := FALSE;
       "Flag Heating Ready" := FALSE;
       "Slof Ready" := FALSE;
       "Flag RS Pneumatic 1 Pusher  Advance" := FALSE;
   END_IF;
END_REGION

REGION Network 7: Check Slof 3 Way
   RUNG wire#powerrail
      Contact( "Machine Running" )
      I_Contact( "Photosensor 6" )
      I_Contact( "Photosensor 7" )
      I_Contact( "Photosensor 8" )
      Contact( "Photosensor 9" )
      I_Contact( "Slof Manual Ready" )
      S_Coil( "Slof Manual Ready" )
   END_RUNG
   // the same network as SCL:
   IF "Machine Running" AND NOT "Photosensor 6" AND NOT "Photosensor 7" AND NOT "Photosensor 8" AND "Photosensor 9" AND NOT "Slof Manual Ready" THEN
       "Slof Manual Ready" := TRUE;
   END_IF;
END_REGION

REGION Network 8: Manual Insert Slof
